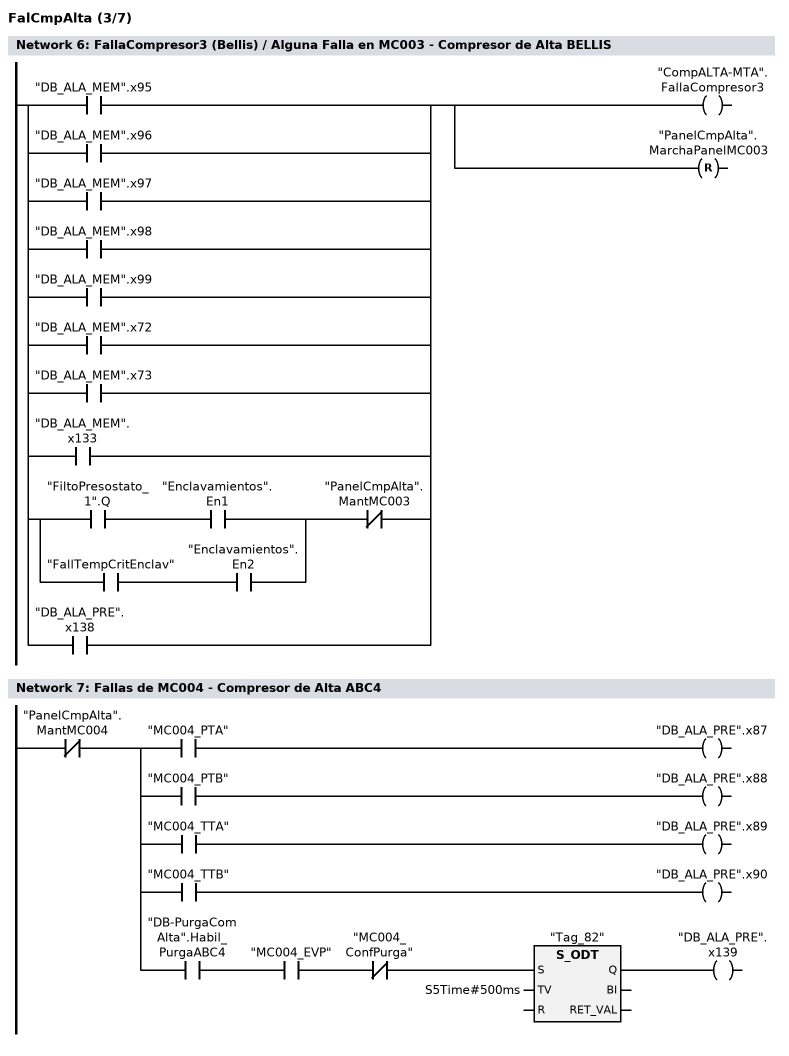
   RUNG wire#powerrail
      Contact( "DB_ALA_MEM".x95 )
      wire#w1
      Coil( "CompALTA-MTA".FallaCompresor3 )
   END_RUNG
   RUNG wire#powerrail
      Contact( "DB_ALA_MEM".x96 )
   END_RUNG wire#w1
   RUNG wire#powerrail
      Contact( "DB_ALA_MEM".x97 )
   END_RUNG wire#w1
   RUNG wire#powerrail
      Contact( "DB_ALA_MEM".x98 )
   END_RUNG wire#w1
   RUNG wire#powerrail
      Contact( "DB_ALA_MEM".x99 )
   END_RUNG wire#w1
   RUNG wire#powerrail
      Contact( "DB_ALA_MEM".x72 )
   END_RUNG wire#w1
   RUNG wire#powerrail
      Contact( "DB_ALA_MEM".x73 )
   END_RUNG wire#w1
   RUNG wire#powerrail
      Contact( "DB_ALA_MEM".x133 )
   END_RUNG wire#w1
   RUNG wire#powerrail
      Contact( "FiltoPresostato_1".Q )
      Contact( "Enclavamientos".En1 )
      wire#w2
      I_Contact( "PanelCmpAlta".MantMC003 )
   END_RUNG wire#w1
   RUNG wire#powerrail
      Contact( "FallTempCritEnclav" )
      Contact( "Enclavamientos".En2 )
   END_RUNG wire#w2
   RUNG wire#powerrail
      Contact( "DB_ALA_PRE".x138 )
   END_RUNG wire#w1
   RUNG wire#w1
      R_Coil( "PanelCmpAlta".MarchaPanelMC003 )
   END_RUNG
   // the same network as SCL:
   "CompALTA-MTA".FallaCompresor3 := "DB_ALA_MEM".x95 OR "DB_ALA_MEM".x96 OR "DB_ALA_MEM".x97 OR "DB_ALA_MEM".x98 OR "DB_ALA_MEM".x99 OR "DB_ALA_MEM".x72 OR "DB_ALA_MEM".x73 OR "DB_ALA_MEM".x133 OR ((("FiltoPresostato_1".Q AND "Enclavamientos".En1) OR ("FallTempCritEnclav" AND "Enclavamientos".En2)) AND NOT "PanelCmpAlta".MantMC003) OR "DB_ALA_PRE".x138;
   IF "CompALTA-MTA".FallaCompresor3 THEN "PanelCmpAlta".MarchaPanelMC003 := FALSE; END_IF;
END_REGION

REGION Network 7: Fallas de MC004 - Compresor de Alta ABC4
   RUNG wire#powerrail
      I_Contact( "PanelCmpAlta".MantMC004 )
      wire#w1
      Contact( "MC004_PTA" )
      Coil( "DB_ALA_PRE".x87 )
   END_RUNG
   RUNG wire#w1
      Contact( "MC004_PTB" )
      Coil( "DB_ALA_PRE".x88 )
   END_RUNG
   RUNG wire#w1
      Contact( "MC004_TTA" )
      Coil( "DB_ALA_PRE".x89 )
   END_RUNG
   RUNG wire#w1
      Contact( "MC004_TTB" )
      Coil( "DB_ALA_PRE".x90 )
   END_RUNG
   RUNG wire#w1
      Contact( "DB-PurgaComAlta".Habil_PurgaABC4 )
      Contact( "MC004_EVP" )
      I_Contact( "MC004_ConfPurga" )
      S_ODT(T_NO := "Tag_82", TV := S5Time#500ms, R :=, BI =>, RET_VAL =>)
      Coil( "DB_ALA_PRE".x139 )
   END_RUNG
   // the same network as SCL:
   #_w1 := NOT "PanelCmpAlta".MantMC004;
   "DB_ALA_PRE".x87 := #_w1 AND "MC004_PTA";
   "DB_ALA_PRE".x88 := #_w1 AND "MC004_PTB";
   "DB_ALA_PRE".x89 := #_w1 AND "MC004_TTA";
   "DB_ALA_PRE".x90 := #_w1 AND "MC004_TTB";
   #_s5time1 := S_ODT(T_NO := "Tag_82",
                      S := #_w1 AND "DB-PurgaComAlta".Habil_PurgaABC4 AND "MC004_EVP" AND NOT "MC004_ConfPurga",
                      TV := S5Time#500ms,
                      Q => #_w2);
   "DB_ALA_PRE".x139 := #_w2;
END_REGION

REGION Network 8: FallaCompresor4 (ABC4) / Alguna Falla en MC004 - Compresor de Alta ABC4
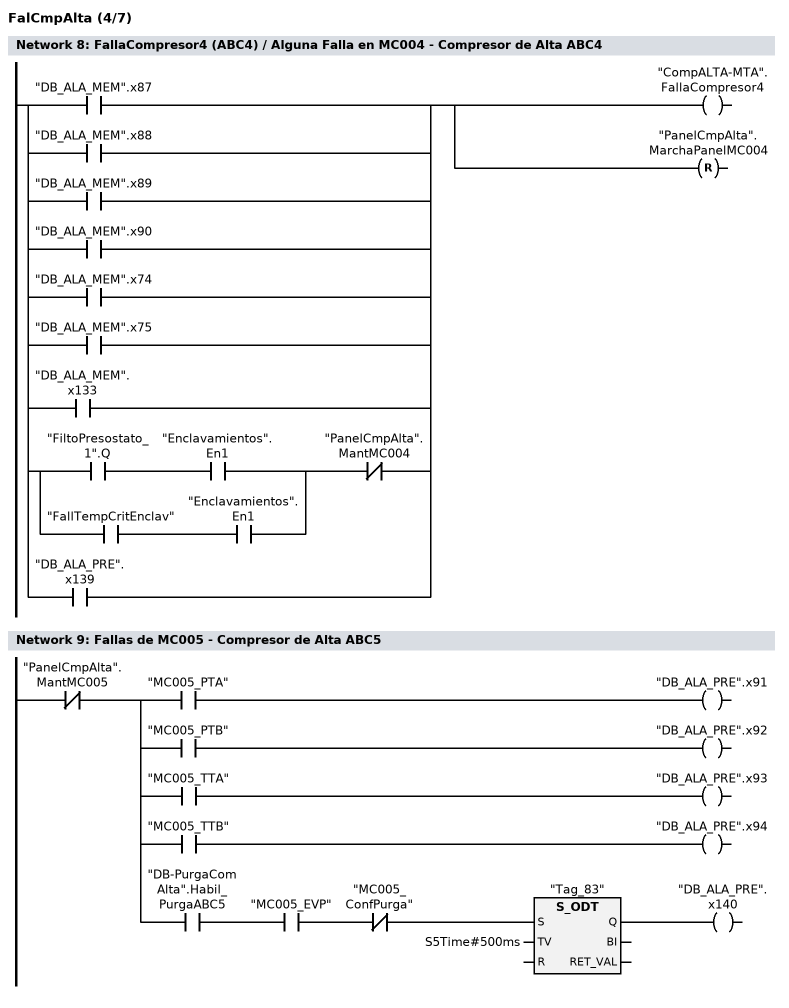
   RUNG wire#powerrail
      Contact( "DB_ALA_MEM".x87 )
      wire#w1
      Coil( "CompALTA-MTA".FallaCompresor4 )
   END_RUNG
   RUNG wire#powerrail
      Contact( "DB_ALA_MEM".x88 )
   END_RUNG wire#w1
   RUNG wire#powerrail
      Contact( "DB_ALA_MEM".x89 )
   END_RUNG wire#w1
   RUNG wire#powerrail
      Contact( "DB_ALA_MEM".x90 )
   END_RUNG wire#w1
   RUNG wire#powerrail
      Contact( "DB_ALA_MEM".x74 )
   END_RUNG wire#w1
   RUNG wire#powerrail
      Contact( "DB_ALA_MEM".x75 )
   END_RUNG wire#w1
   RUNG wire#powerrail
      Contact( "DB_ALA_MEM".x133 )
   END_RUNG wire#w1
   RUNG wire#powerrail
      Contact( "FiltoPresostato_1".Q )
      Contact( "Enclavamientos".En1 )
      wire#w2
      I_Contact( "PanelCmpAlta".MantMC004 )
   END_RUNG wire#w1
   RUNG wire#powerrail
      Contact( "FallTempCritEnclav" )
      Contact( "Enclavamientos".En1 )
   END_RUNG wire#w2
   RUNG wire#powerrail
      Contact( "DB_ALA_PRE".x139 )
   END_RUNG wire#w1
   RUNG wire#w1
      R_Coil( "PanelCmpAlta".MarchaPanelMC004 )
   END_RUNG
   // the same network as SCL:
   "CompALTA-MTA".FallaCompresor4 := "DB_ALA_MEM".x87 OR "DB_ALA_MEM".x88 OR "DB_ALA_MEM".x89 OR "DB_ALA_MEM".x90 OR "DB_ALA_MEM".x74 OR "DB_ALA_MEM".x75 OR "DB_ALA_MEM".x133 OR ((("FiltoPresostato_1".Q AND "Enclavamientos".En1) OR ("FallTempCritEnclav" AND "Enclavamientos".En1)) AND NOT "PanelCmpAlta".MantMC004) OR "DB_ALA_PRE".x139;
   IF "CompALTA-MTA".FallaCompresor4 THEN "PanelCmpAlta".MarchaPanelMC004 := FALSE; END_IF;
END_REGION

REGION Network 9: Fallas de MC005 - Compresor de Alta ABC5
   RUNG wire#powerrail
      I_Contact( "PanelCmpAlta".MantMC005 )
      wire#w1
      Contact( "MC005_PTA" )
      Coil( "DB_ALA_PRE".x91 )
   END_RUNG
   RUNG wire#w1
      Contact( "MC005_PTB" )
      Coil( "DB_ALA_PRE".x92 )
   END_RUNG
   RUNG wire#w1
      Contact( "MC005_TTA" )
      Coil( "DB_ALA_PRE".x93 )
   END_RUNG
   RUNG wire#w1
      Contact( "MC005_TTB" )
      Coil( "DB_ALA_PRE".x94 )
   END_RUNG
   RUNG wire#w1
      Contact( "DB-PurgaComAlta".Habil_PurgaABC5 )
      Contact( "MC005_EVP" )
      I_Contact( "MC005_ConfPurga" )
      S_ODT(T_NO := "Tag_83", TV := S5Time#500ms, R :=, BI =>, RET_VAL =>)
      Coil( "DB_ALA_PRE".x140 )
   END_RUNG
   // the same network as SCL:
   #_w1 := NOT "PanelCmpAlta".MantMC005;
   "DB_ALA_PRE".x91 := #_w1 AND "MC005_PTA";
   "DB_ALA_PRE".x92 := #_w1 AND "MC005_PTB";
   "DB_ALA_PRE".x93 := #_w1 AND "MC005_TTA";
   "DB_ALA_PRE".x94 := #_w1 AND "MC005_TTB";
   #_s5time1 := S_ODT(T_NO := "Tag_83",
                      S := #_w1 AND "DB-PurgaComAlta".Habil_PurgaABC5 AND "MC005_EVP" AND NOT "MC005_ConfPurga",
                      TV := S5Time#500ms,
                      Q => #_w2);
   "DB_ALA_PRE".x140 := #_w2;
END_REGION

REGION Network 10: FallaCompresor5 (ABC5) / Alguna Falla en MC005 - Compresor de Alta ABC5
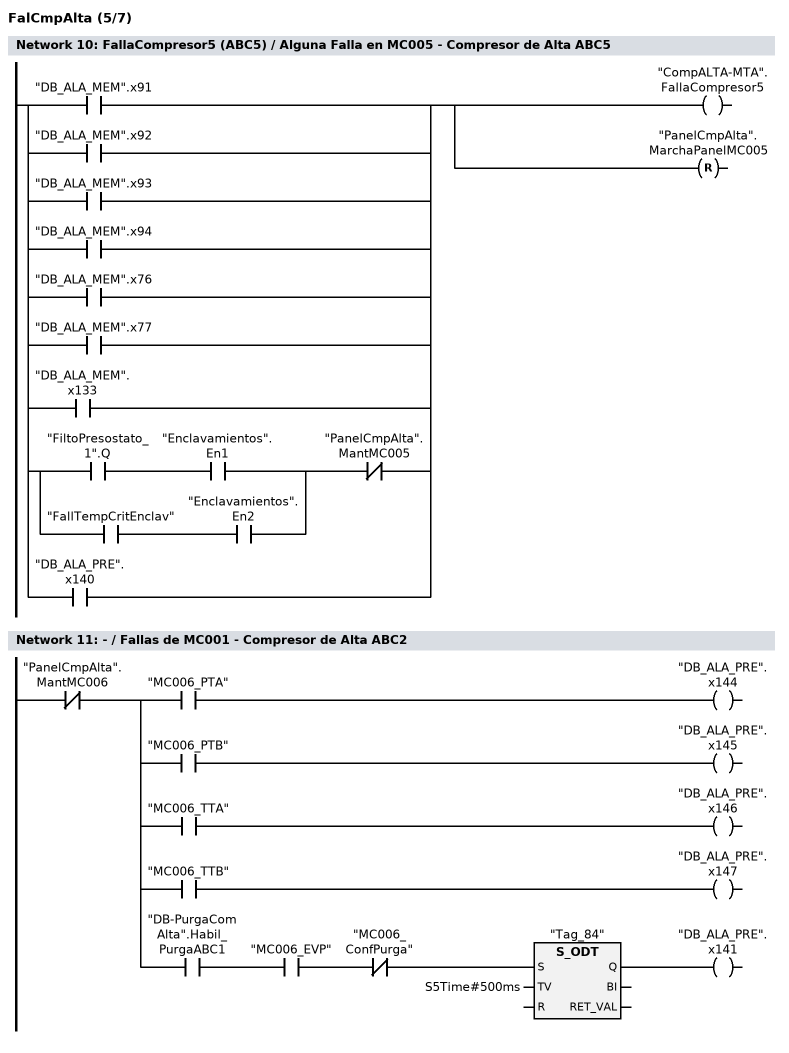
   RUNG wire#powerrail
      Contact( "DB_ALA_MEM".x91 )
      wire#w1
      Coil( "CompALTA-MTA".FallaCompresor5 )
   END_RUNG
   RUNG wire#powerrail
      Contact( "DB_ALA_MEM".x92 )
   END_RUNG wire#w1
   RUNG wire#powerrail
      Contact( "DB_ALA_MEM".x93 )
   END_RUNG wire#w1
   RUNG wire#powerrail
      Contact( "DB_ALA_MEM".x94 )
   END_RUNG wire#w1
   RUNG wire#powerrail
      Contact( "DB_ALA_MEM".x76 )
   END_RUNG wire#w1
   RUNG wire#powerrail
      Contact( "DB_ALA_MEM".x77 )
   END_RUNG wire#w1
   RUNG wire#powerrail
      Contact( "DB_ALA_MEM".x133 )
   END_RUNG wire#w1
   RUNG wire#powerrail
      Contact( "FiltoPresostato_1".Q )
      Contact( "Enclavamientos".En1 )
      wire#w2
      I_Contact( "PanelCmpAlta".MantMC005 )
   END_RUNG wire#w1
   RUNG wire#powerrail
      Contact( "FallTempCritEnclav" )
      Contact( "Enclavamientos".En2 )
   END_RUNG wire#w2
   RUNG wire#powerrail
      Contact( "DB_ALA_PRE".x140 )
   END_RUNG wire#w1
   RUNG wire#w1
      R_Coil( "PanelCmpAlta".MarchaPanelMC005 )
   END_RUNG
   // the same network as SCL:
   "CompALTA-MTA".FallaCompresor5 := "DB_ALA_MEM".x91 OR "DB_ALA_MEM".x92 OR "DB_ALA_MEM".x93 OR "DB_ALA_MEM".x94 OR "DB_ALA_MEM".x76 OR "DB_ALA_MEM".x77 OR "DB_ALA_MEM".x133 OR ((("FiltoPresostato_1".Q AND "Enclavamientos".En1) OR ("FallTempCritEnclav" AND "Enclavamientos".En2)) AND NOT "PanelCmpAlta".MantMC005) OR "DB_ALA_PRE".x140;
   IF "CompALTA-MTA".FallaCompresor5 THEN "PanelCmpAlta".MarchaPanelMC005 := FALSE; END_IF;
END_REGION

REGION Network 11: - / Fallas de MC001 - Compresor de Alta ABC2
   RUNG wire#powerrail
      I_Contact( "PanelCmpAlta".MantMC006 )
      wire#w1
      Contact( "MC006_PTA" )
      Coil( "DB_ALA_PRE".x144 )
   END_RUNG
   RUNG wire#w1
      Contact( "MC006_PTB" )
      Coil( "DB_ALA_PRE".x145 )
   END_RUNG
   RUNG wire#w1
      Contact( "MC006_TTA" )
      Coil( "DB_ALA_PRE".x146 )
   END_RUNG
   RUNG wire#w1
      Contact( "MC006_TTB" )
      Coil( "DB_ALA_PRE".x147 )
   END_RUNG
   RUNG wire#w1
      Contact( "DB-PurgaComAlta".Habil_PurgaABC1 )
      Contact( "MC006_EVP" )
      I_Contact( "MC006_ConfPurga" )
      S_ODT(T_NO := "Tag_84", TV := S5Time#500ms, R :=, BI =>, RET_VAL =>)
      Coil( "DB_ALA_PRE".x141 )
   END_RUNG
   // the same network as SCL:
   #_w1 := NOT "PanelCmpAlta".MantMC006;
   "DB_ALA_PRE".x144 := #_w1 AND "MC006_PTA";
   "DB_ALA_PRE".x145 := #_w1 AND "MC006_PTB";
   "DB_ALA_PRE".x146 := #_w1 AND "MC006_TTA";
   "DB_ALA_PRE".x147 := #_w1 AND "MC006_TTB";
   #_s5time1 := S_ODT(T_NO := "Tag_84",
                      S := #_w1 AND "DB-PurgaComAlta".Habil_PurgaABC1 AND "MC006_EVP" AND NOT "MC006_ConfPurga",
                      TV := S5Time#500ms,
                      Q => #_w2);
   "DB_ALA_PRE".x141 := #_w2;
END_REGION

REGION Network 12: FallaCompresor6 (ABC1) / Alguna Falla en MC001 - Compresor de Alta ABC2
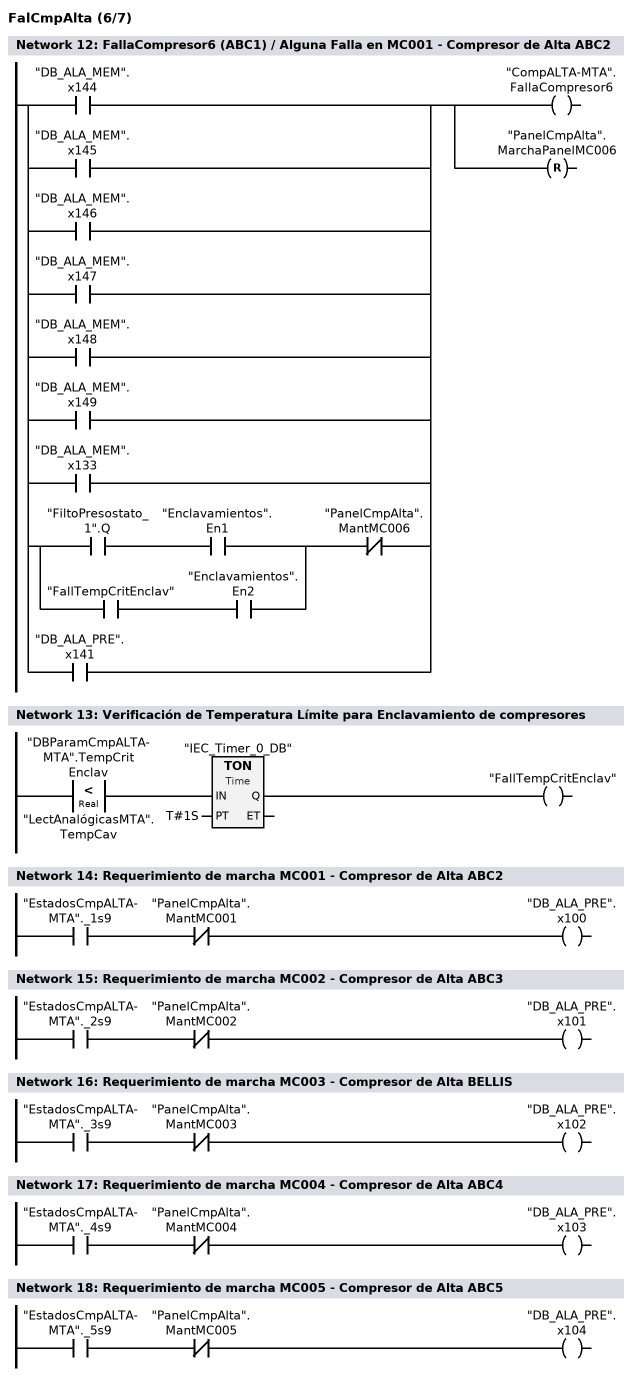
   RUNG wire#powerrail
      Contact( "DB_ALA_MEM".x144 )
      wire#w1
      Coil( "CompALTA-MTA".FallaCompresor6 )
   END_RUNG
   RUNG wire#powerrail
      Contact( "DB_ALA_MEM".x145 )
   END_RUNG wire#w1
   RUNG wire#powerrail
      Contact( "DB_ALA_MEM".x146 )
   END_RUNG wire#w1
   RUNG wire#powerrail
      Contact( "DB_ALA_MEM".x147 )
   END_RUNG wire#w1
   RUNG wire#powerrail
      Contact( "DB_ALA_MEM".x148 )
   END_RUNG wire#w1
   RUNG wire#powerrail
      Contact( "DB_ALA_MEM".x149 )
   END_RUNG wire#w1
   RUNG wire#powerrail
      Contact( "DB_ALA_MEM".x133 )
   END_RUNG wire#w1
   RUNG wire#powerrail
      Contact( "FiltoPresostato_1".Q )
      Contact( "Enclavamientos".En1 )
      wire#w2
      I_Contact( "PanelCmpAlta".MantMC006 )
   END_RUNG wire#w1
   RUNG wire#powerrail
      Contact( "FallTempCritEnclav" )
      Contact( "Enclavamientos".En2 )
   END_RUNG wire#w2
   RUNG wire#powerrail
      Contact( "DB_ALA_PRE".x141 )
   END_RUNG wire#w1
   RUNG wire#w1
      R_Coil( "PanelCmpAlta".MarchaPanelMC006 )
   END_RUNG
   // the same network as SCL:
   "CompALTA-MTA".FallaCompresor6 := "DB_ALA_MEM".x144 OR "DB_ALA_MEM".x145 OR "DB_ALA_MEM".x146 OR "DB_ALA_MEM".x147 OR "DB_ALA_MEM".x148 OR "DB_ALA_MEM".x149 OR "DB_ALA_MEM".x133 OR ((("FiltoPresostato_1".Q AND "Enclavamientos".En1) OR ("FallTempCritEnclav" AND "Enclavamientos".En2)) AND NOT "PanelCmpAlta".MantMC006) OR "DB_ALA_PRE".x141;
   IF "CompALTA-MTA".FallaCompresor6 THEN "PanelCmpAlta".MarchaPanelMC006 := FALSE; END_IF;
END_REGION

REGION Network 13: Verificación de Temperatura Límite para Enclavamiento de compresores
   "IEC_Timer_0_DB".TON(IN := "DBParamCmpALTA-MTA".TempCritEnclav < "LectAnalógicasMTA".TempCav, PT := T#1S);
   "FallTempCritEnclav" := "IEC_Timer_0_DB".Q;
END_REGION

REGION Network 14: Requerimiento de marcha MC001 - Compresor de Alta ABC2
   RUNG wire#powerrail
      Contact( "EstadosCmpALTA-MTA"._1s9 )
      I_Contact( "PanelCmpAlta".MantMC001 )
      Coil( "DB_ALA_PRE".x100 )
   END_RUNG
   // the same network as SCL:
   "DB_ALA_PRE".x100 := "EstadosCmpALTA-MTA"._1s9 AND NOT "PanelCmpAlta".MantMC001;
END_REGION

REGION Network 15: Requerimiento de marcha MC002 - Compresor de Alta ABC3
   RUNG wire#powerrail
      Contact( "EstadosCmpALTA-MTA"._2s9 )
      I_Contact( "PanelCmpAlta".MantMC002 )
      Coil( "DB_ALA_PRE".x101 )
   END_RUNG
   // the same network as SCL:
   "DB_ALA_PRE".x101 := "EstadosCmpALTA-MTA"._2s9 AND NOT "PanelCmpAlta".MantMC002;
END_REGION

REGION Network 16: Requerimiento de marcha MC003 - Compresor de Alta BELLIS
   RUNG wire#powerrail
      Contact( "EstadosCmpALTA-MTA"._3s9 )
      I_Contact( "PanelCmpAlta".MantMC003 )
      Coil( "DB_ALA_PRE".x102 )
   END_RUNG
   // the same network as SCL:
   "DB_ALA_PRE".x102 := "EstadosCmpALTA-MTA"._3s9 AND NOT "PanelCmpAlta".MantMC003;
END_REGION

REGION Network 17: Requerimiento de marcha MC004 - Compresor de Alta ABC4
   RUNG wire#powerrail
      Contact( "EstadosCmpALTA-MTA"._4s9 )
      I_Contact( "PanelCmpAlta".MantMC004 )
      Coil( "DB_ALA_PRE".x103 )
   END_RUNG
   // the same network as SCL:
   "DB_ALA_PRE".x103 := "EstadosCmpALTA-MTA"._4s9 AND NOT "PanelCmpAlta".MantMC004;
END_REGION

REGION Network 18: Requerimiento de marcha MC005 - Compresor de Alta ABC5
   RUNG wire#powerrail
      Contact( "EstadosCmpALTA-MTA"._5s9 )
      I_Contact( "PanelCmpAlta".MantMC005 )
      Coil( "DB_ALA_PRE".x104 )
   END_RUNG
   // the same network as SCL:
   "DB_ALA_PRE".x104 := "EstadosCmpALTA-MTA"._5s9 AND NOT "PanelCmpAlta".MantMC005;
END_REGION

REGION Network 19: Requerimiento de marcha MC001 - Compresor de Alta ABC2
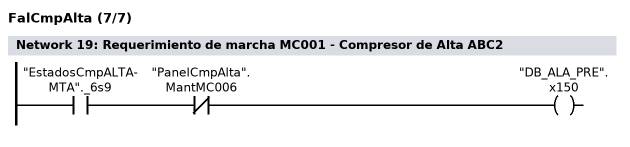
   RUNG wire#powerrail
      Contact( "EstadosCmpALTA-MTA"._6s9 )
      I_Contact( "PanelCmpAlta".MantMC006 )
      Coil( "DB_ALA_PRE".x150 )
   END_RUNG
   // the same network as SCL:
   "DB_ALA_PRE".x150 := "EstadosCmpALTA-MTA"._6s9 AND NOT "PanelCmpAlta".MantMC006;
END_REGION
END_FUNCTION

// folder: Auxiliares

FUNCTION "AjusteEntrada-SalidaMTA" : Void   // FC6, LAD
{ S7_Optimized_Access := 'FALSE' }
VERSION : 0.1
BEGIN

REGION Network 1
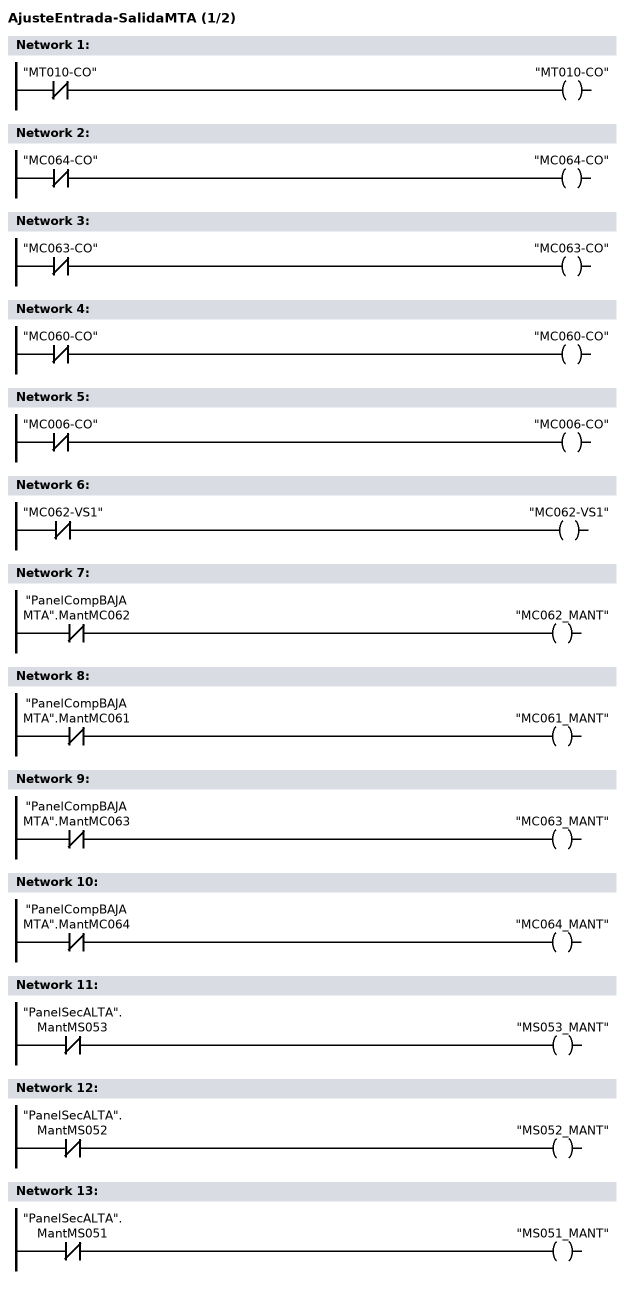
   RUNG wire#powerrail
      I_Contact( "MT010-CO" )
      Coil( "MT010-CO" )
   END_RUNG
   // the same network as SCL:
   "MT010-CO" := NOT "MT010-CO";
END_REGION

REGION Network 2
   RUNG wire#powerrail
      I_Contact( "MC064-CO" )
      Coil( "MC064-CO" )
   END_RUNG
   // the same network as SCL:
   "MC064-CO" := NOT "MC064-CO";
END_REGION

REGION Network 3
   RUNG wire#powerrail
      I_Contact( "MC063-CO" )
      Coil( "MC063-CO" )
   END_RUNG
   // the same network as SCL:
   "MC063-CO" := NOT "MC063-CO";
END_REGION

REGION Network 4
   RUNG wire#powerrail
      I_Contact( "MC060-CO" )
      Coil( "MC060-CO" )
   END_RUNG
   // the same network as SCL:
   "MC060-CO" := NOT "MC060-CO";
END_REGION

REGION Network 5
   RUNG wire#powerrail
      I_Contact( "MC006-CO" )
      Coil( "MC006-CO" )
   END_RUNG
   // the same network as SCL:
   "MC006-CO" := NOT "MC006-CO";
END_REGION

REGION Network 6
   RUNG wire#powerrail
      I_Contact( "MC062-VS1" )
      Coil( "MC062-VS1" )
   END_RUNG
   // the same network as SCL:
   "MC062-VS1" := NOT "MC062-VS1";
END_REGION

REGION Network 7
   RUNG wire#powerrail
      I_Contact( "PanelCompBAJA MTA".MantMC062 )
      Coil( "MC062_MANT" )
   END_RUNG
   // the same network as SCL:
   "MC062_MANT" := NOT "PanelCompBAJA MTA".MantMC062;
END_REGION

REGION Network 8
   RUNG wire#powerrail
      I_Contact( "PanelCompBAJA MTA".MantMC061 )
      Coil( "MC061_MANT" )
   END_RUNG
   // the same network as SCL:
   "MC061_MANT" := NOT "PanelCompBAJA MTA".MantMC061;
END_REGION

REGION Network 9
   RUNG wire#powerrail
      I_Contact( "PanelCompBAJA MTA".MantMC063 )
      Coil( "MC063_MANT" )
   END_RUNG
   // the same network as SCL:
   "MC063_MANT" := NOT "PanelCompBAJA MTA".MantMC063;
END_REGION

REGION Network 10
   RUNG wire#powerrail
      I_Contact( "PanelCompBAJA MTA".MantMC064 )
      Coil( "MC064_MANT" )
   END_RUNG
   // the same network as SCL:
   "MC064_MANT" := NOT "PanelCompBAJA MTA".MantMC064;
END_REGION

REGION Network 11
   RUNG wire#powerrail
      I_Contact( "PanelSecALTA".MantMS053 )
      Coil( "MS053_MANT" )
   END_RUNG
   // the same network as SCL:
   "MS053_MANT" := NOT "PanelSecALTA".MantMS053;
END_REGION

REGION Network 12
   RUNG wire#powerrail
      I_Contact( "PanelSecALTA".MantMS052 )
      Coil( "MS052_MANT" )
   END_RUNG
   // the same network as SCL:
   "MS052_MANT" := NOT "PanelSecALTA".MantMS052;
END_REGION

REGION Network 13
   RUNG wire#powerrail
      I_Contact( "PanelSecALTA".MantMS051 )
      Coil( "MS051_MANT" )
   END_RUNG
   // the same network as SCL:
   "MS051_MANT" := NOT "PanelSecALTA".MantMS051;
END_REGION

REGION Network 14
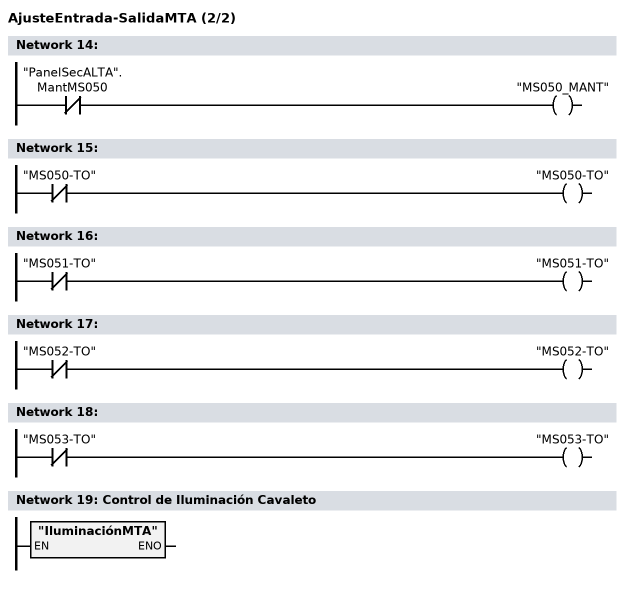
   RUNG wire#powerrail
      I_Contact( "PanelSecALTA".MantMS050 )
      Coil( "MS050_MANT" )
   END_RUNG
   // the same network as SCL:
   "MS050_MANT" := NOT "PanelSecALTA".MantMS050;
END_REGION

REGION Network 15
   RUNG wire#powerrail
      I_Contact( "MS050-TO" )
      Coil( "MS050-TO" )
   END_RUNG
   // the same network as SCL:
   "MS050-TO" := NOT "MS050-TO";
END_REGION

REGION Network 16
   RUNG wire#powerrail
      I_Contact( "MS051-TO" )
      Coil( "MS051-TO" )
   END_RUNG
   // the same network as SCL:
   "MS051-TO" := NOT "MS051-TO";
END_REGION

REGION Network 17
   RUNG wire#powerrail
      I_Contact( "MS052-TO" )
      Coil( "MS052-TO" )
   END_RUNG
   // the same network as SCL:
   "MS052-TO" := NOT "MS052-TO";
END_REGION

REGION Network 18
   RUNG wire#powerrail
      I_Contact( "MS053-TO" )
      Coil( "MS053-TO" )
   END_RUNG
   // the same network as SCL:
   "MS053-TO" := NOT "MS053-TO";
END_REGION

REGION Network 19: Control de Iluminación Cavaleto
   RUNG wire#powerrail
      "IluminaciónMTA"()
   END_RUNG
   // the same network as SCL:
   "IluminaciónMTA"();
END_REGION
END_FUNCTION

FUNCTION "And-Byte MTA" : Void   // FC22, LAD
{ S7_Optimized_Access := 'FALSE' }
VERSION : 0.1
BEGIN

REGION Network 1
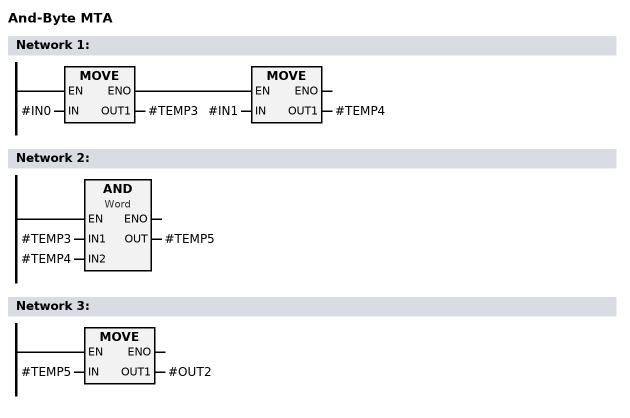
   RUNG wire#powerrail
      { S7_GenerateENO := "TRUE" } Move(in := #IN0, out1 => #TEMP3)
      { S7_GenerateENO := "TRUE" } Move(in := #IN1, out1 => #TEMP4)
   END_RUNG
   // the same network as SCL:
   // ENO of a box is taken as its EN; it also drops when the box reports an error
   #TEMP3 := #IN0;
   #TEMP4 := #IN1;
END_REGION

REGION Network 2
   RUNG wire#powerrail
      { S7_Templates := "SrcType := Word"; S7_GenerateENO := "TRUE" } And(in1 := #TEMP3, in2 := #TEMP4, out => #TEMP5)
   END_RUNG
   // the same network as SCL:
   #TEMP5 := #TEMP3 AND #TEMP4;
END_REGION

REGION Network 3
   RUNG wire#powerrail
      { S7_GenerateENO := "TRUE" } Move(in := #TEMP5, out1 => #OUT2)
   END_RUNG
   // the same network as SCL:
   #OUT2 := #TEMP5;
END_REGION
END_FUNCTION

FUNCTION "Inicialización" : Void   // FC46, LAD
{ S7_Optimized_Access := 'FALSE' }
VERSION : 0.1
BEGIN

REGION Network 1
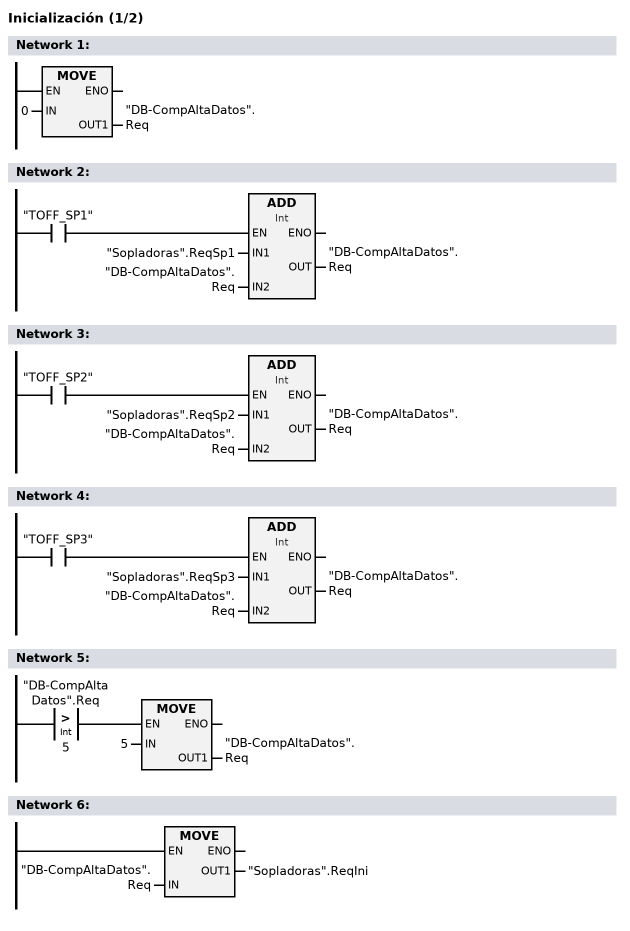
   RUNG wire#powerrail
      { S7_GenerateENO := "TRUE" } Move(in := 0, out1 => "DB-CompAltaDatos".Req)
   END_RUNG
   // the same network as SCL:
   "DB-CompAltaDatos".Req := 0;
END_REGION

REGION Network 2
   RUNG wire#powerrail
      Contact( "TOFF_SP1" )
      { S7_Templates := "SrcType := Int"; S7_GenerateENO := "TRUE" } Add(in1 := "Sopladoras".ReqSp1, in2 := "DB-CompAltaDatos".Req, out => "DB-CompAltaDatos".Req)
   END_RUNG
   // the same network as SCL:
   IF "TOFF_SP1" THEN "DB-CompAltaDatos".Req := "Sopladoras".ReqSp1 + "DB-CompAltaDatos".Req; END_IF;
END_REGION

REGION Network 3
   RUNG wire#powerrail
      Contact( "TOFF_SP2" )
      { S7_Templates := "SrcType := Int"; S7_GenerateENO := "TRUE" } Add(in1 := "Sopladoras".ReqSp2, in2 := "DB-CompAltaDatos".Req, out => "DB-CompAltaDatos".Req)
   END_RUNG
   // the same network as SCL:
   IF "TOFF_SP2" THEN "DB-CompAltaDatos".Req := "Sopladoras".ReqSp2 + "DB-CompAltaDatos".Req; END_IF;
END_REGION

REGION Network 4
   RUNG wire#powerrail
      Contact( "TOFF_SP3" )
      { S7_Templates := "SrcType := Int"; S7_GenerateENO := "TRUE" } Add(in1 := "Sopladoras".ReqSp3, in2 := "DB-CompAltaDatos".Req, out => "DB-CompAltaDatos".Req)
   END_RUNG
   // the same network as SCL:
   IF "TOFF_SP3" THEN "DB-CompAltaDatos".Req := "Sopladoras".ReqSp3 + "DB-CompAltaDatos".Req; END_IF;
END_REGION

REGION Network 5
   RUNG wire#powerrail
      { S7_Templates := "SrcType := Int" } GT_Contact(in1 := "DB-CompAltaDatos".Req, in2 := 5)
      { S7_GenerateENO := "TRUE" } Move(in := 5, out1 => "DB-CompAltaDatos".Req)
   END_RUNG
   // the same network as SCL:
   IF "DB-CompAltaDatos".Req > 5 THEN "DB-CompAltaDatos".Req := 5; END_IF;
END_REGION

REGION Network 6
   RUNG wire#powerrail
      { S7_GenerateENO := "TRUE" } Move(in := "DB-CompAltaDatos".Req, out1 => "Sopladoras".ReqIni)
   END_RUNG
   // the same network as SCL:
   "Sopladoras".ReqIni := "DB-CompAltaDatos".Req;
END_REGION

REGION Network 7
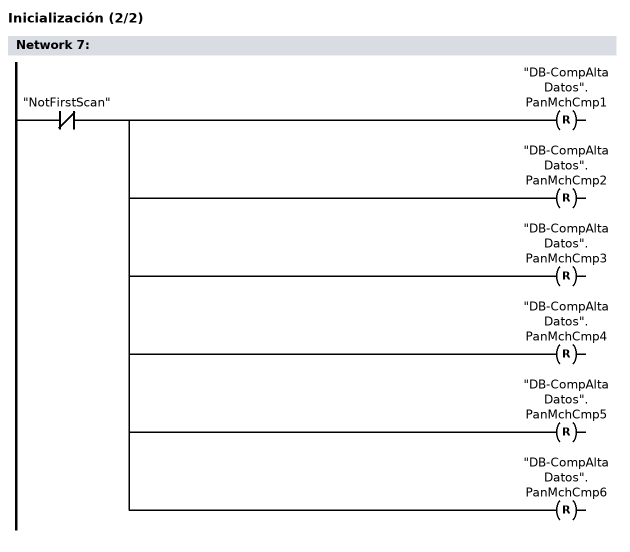
   RUNG wire#powerrail
      I_Contact( "NotFirstScan" )
      wire#w1
      R_Coil( "DB-CompAltaDatos".PanMchCmp1 )
   END_RUNG
   RUNG wire#w1
      R_Coil( "DB-CompAltaDatos".PanMchCmp2 )
   END_RUNG
   RUNG wire#w1
      R_Coil( "DB-CompAltaDatos".PanMchCmp3 )
   END_RUNG
   RUNG wire#w1
      R_Coil( "DB-CompAltaDatos".PanMchCmp4 )
   END_RUNG
   RUNG wire#w1
      R_Coil( "DB-CompAltaDatos".PanMchCmp5 )
   END_RUNG
   RUNG wire#w1
      R_Coil( "DB-CompAltaDatos".PanMchCmp6 )
   END_RUNG
   // the same network as SCL:
   IF NOT "NotFirstScan" THEN
       "DB-CompAltaDatos".PanMchCmp1 := FALSE;
       "DB-CompAltaDatos".PanMchCmp2 := FALSE;
       "DB-CompAltaDatos".PanMchCmp3 := FALSE;
       "DB-CompAltaDatos".PanMchCmp4 := FALSE;
       "DB-CompAltaDatos".PanMchCmp5 := FALSE;
       "DB-CompAltaDatos".PanMchCmp6 := FALSE;
   END_IF;
END_REGION
END_FUNCTION

// folder: Bloques Estándar

FUNCTION_BLOCK "ControladorMotoresMTA"   // FB2, LAD
{ S7_Optimized_Access := 'FALSE' }
VERSION : 0.1
BEGIN

REGION Network 2
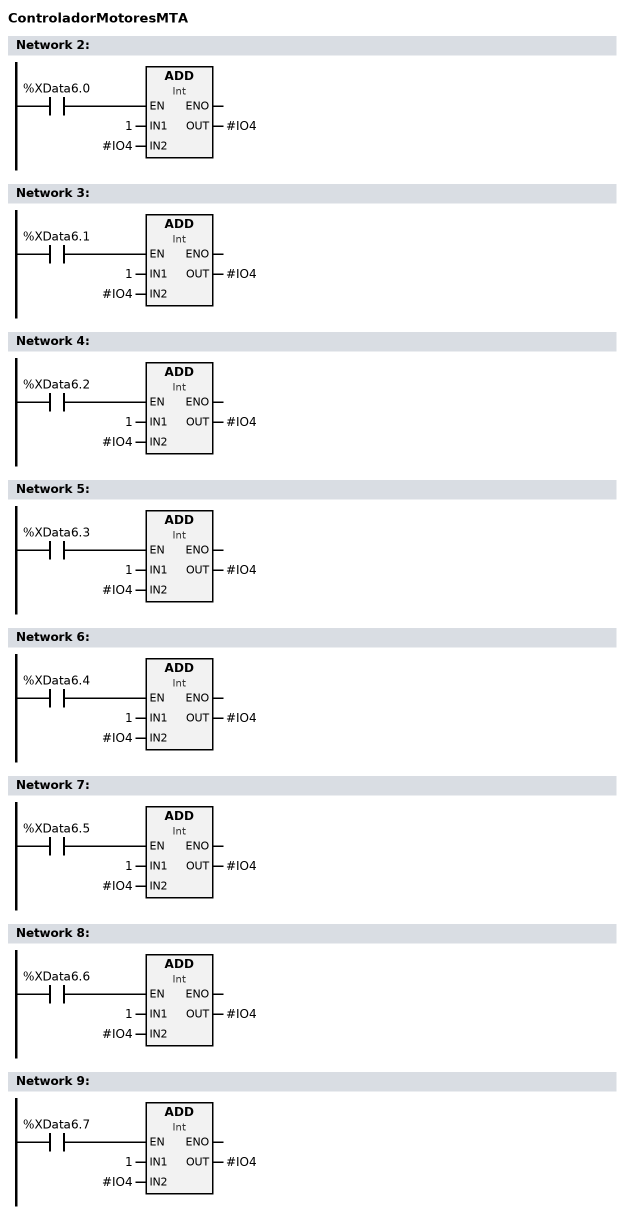
   RUNG wire#powerrail
      Contact( %XData6.0 )
      { S7_Templates := "SrcType := Int"; S7_GenerateENO := "TRUE" } Add(in1 := 1, in2 := #IO4, out => #IO4)
   END_RUNG
   // the same network as SCL:
   IF %XData6.0 THEN #IO4 := 1 + #IO4; END_IF;
END_REGION

REGION Network 3
   RUNG wire#powerrail
      Contact( %XData6.1 )
      { S7_Templates := "SrcType := Int"; S7_GenerateENO := "TRUE" } Add(in1 := 1, in2 := #IO4, out => #IO4)
   END_RUNG
   // the same network as SCL:
   IF %XData6.1 THEN #IO4 := 1 + #IO4; END_IF;
END_REGION

REGION Network 4
   RUNG wire#powerrail
      Contact( %XData6.2 )
      { S7_Templates := "SrcType := Int"; S7_GenerateENO := "TRUE" } Add(in1 := 1, in2 := #IO4, out => #IO4)
   END_RUNG
   // the same network as SCL:
   IF %XData6.2 THEN #IO4 := 1 + #IO4; END_IF;
END_REGION

REGION Network 5
   RUNG wire#powerrail
      Contact( %XData6.3 )
      { S7_Templates := "SrcType := Int"; S7_GenerateENO := "TRUE" } Add(in1 := 1, in2 := #IO4, out => #IO4)
   END_RUNG
   // the same network as SCL:
   IF %XData6.3 THEN #IO4 := 1 + #IO4; END_IF;
END_REGION

REGION Network 6
   RUNG wire#powerrail
      Contact( %XData6.4 )
      { S7_Templates := "SrcType := Int"; S7_GenerateENO := "TRUE" } Add(in1 := 1, in2 := #IO4, out => #IO4)
   END_RUNG
   // the same network as SCL:
   IF %XData6.4 THEN #IO4 := 1 + #IO4; END_IF;
END_REGION

REGION Network 7
   RUNG wire#powerrail
      Contact( %XData6.5 )
      { S7_Templates := "SrcType := Int"; S7_GenerateENO := "TRUE" } Add(in1 := 1, in2 := #IO4, out => #IO4)
   END_RUNG
   // the same network as SCL:
   IF %XData6.5 THEN #IO4 := 1 + #IO4; END_IF;
END_REGION

REGION Network 8
   RUNG wire#powerrail
      Contact( %XData6.6 )
      { S7_Templates := "SrcType := Int"; S7_GenerateENO := "TRUE" } Add(in1 := 1, in2 := #IO4, out => #IO4)
   END_RUNG
   // the same network as SCL:
   IF %XData6.6 THEN #IO4 := 1 + #IO4; END_IF;
END_REGION

REGION Network 9
   RUNG wire#powerrail
      Contact( %XData6.7 )
      { S7_Templates := "SrcType := Int"; S7_GenerateENO := "TRUE" } Add(in1 := 1, in2 := #IO4, out => #IO4)
   END_RUNG
   // the same network as SCL:
   IF %XData6.7 THEN #IO4 := 1 + #IO4; END_IF;
END_REGION
END_FUNCTION_BLOCK

// folder: Compresores/Alta

FUNCTION "CompresoresAltaMTA" : Void   // FC13, LAD
{ S7_Optimized_Access := 'FALSE' }
VERSION : 0.1
BEGIN

REGION Network 1
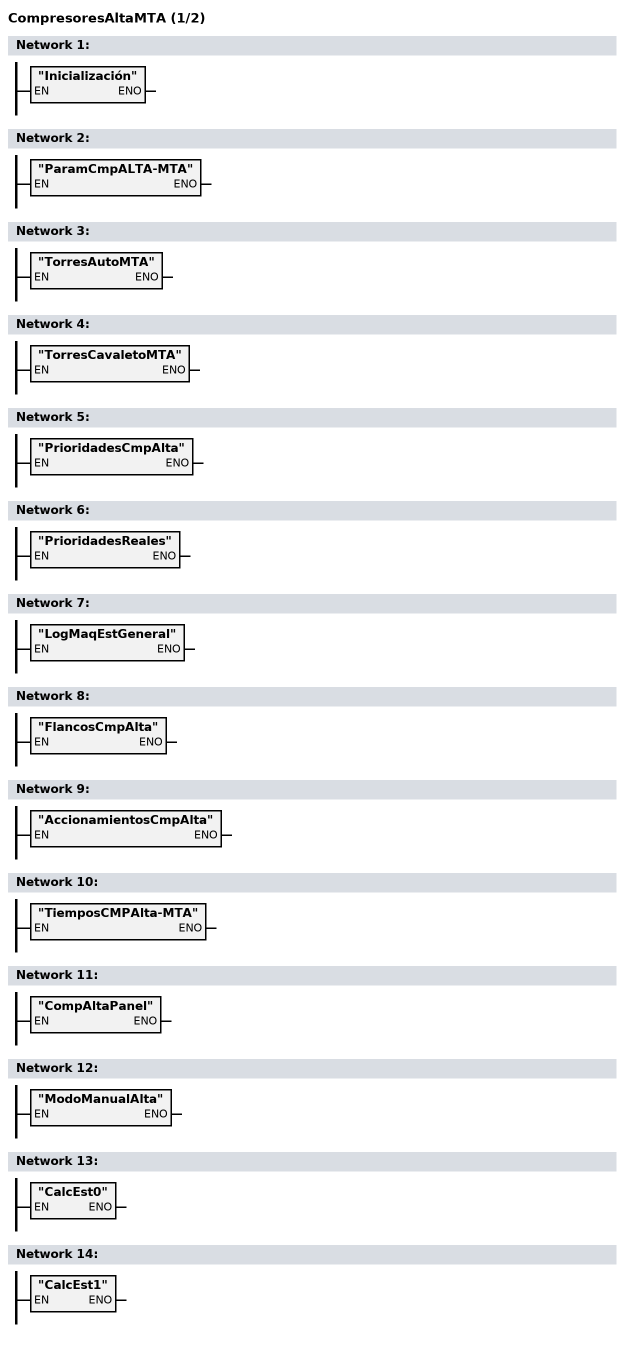
   RUNG wire#powerrail
      "Inicialización"()
   END_RUNG
   // the same network as SCL:
   "Inicialización"();
END_REGION

REGION Network 2
   RUNG wire#powerrail
      "ParamCmpALTA-MTA"()
   END_RUNG
   // the same network as SCL:
   "ParamCmpALTA-MTA"();
END_REGION

REGION Network 3
   RUNG wire#powerrail
      "TorresAutoMTA"()
   END_RUNG
   // the same network as SCL:
   "TorresAutoMTA"();
END_REGION

REGION Network 4
   RUNG wire#powerrail
      "TorresCavaletoMTA"()
   END_RUNG
   // the same network as SCL:
   "TorresCavaletoMTA"();
END_REGION

REGION Network 5
   RUNG wire#powerrail
      "PrioridadesCmpAlta"()
   END_RUNG
   // the same network as SCL:
   "PrioridadesCmpAlta"();
END_REGION

REGION Network 6
   RUNG wire#powerrail
      "PrioridadesReales"()
   END_RUNG
   // the same network as SCL:
   "PrioridadesReales"();
END_REGION

REGION Network 7
   RUNG wire#powerrail
      "LogMaqEstGeneral"()
   END_RUNG
   // the same network as SCL:
   "LogMaqEstGeneral"();
END_REGION

REGION Network 8
   RUNG wire#powerrail
      "FlancosCmpAlta"()
   END_RUNG
   // the same network as SCL:
   "FlancosCmpAlta"();
END_REGION

REGION Network 9
   RUNG wire#powerrail
      "AccionamientosCmpAlta"()
   END_RUNG
   // the same network as SCL:
   "AccionamientosCmpAlta"();
END_REGION

REGION Network 10
   RUNG wire#powerrail
      "TiemposCMPAlta-MTA"()
   END_RUNG
   // the same network as SCL:
   "TiemposCMPAlta-MTA"();
END_REGION

REGION Network 11
   RUNG wire#powerrail
      "CompAltaPanel"()
   END_RUNG
   // the same network as SCL:
   "CompAltaPanel"();
END_REGION

REGION Network 12
   RUNG wire#powerrail
      "ModoManualAlta"()
   END_RUNG
   // the same network as SCL:
   "ModoManualAlta"();
END_REGION

REGION Network 13
   RUNG wire#powerrail
      "CalcEst0"()
   END_RUNG
   // the same network as SCL:
   "CalcEst0"();
END_REGION

REGION Network 14
   RUNG wire#powerrail
      "CalcEst1"()
   END_RUNG
   // the same network as SCL:
   "CalcEst1"();
END_REGION

REGION Network 15
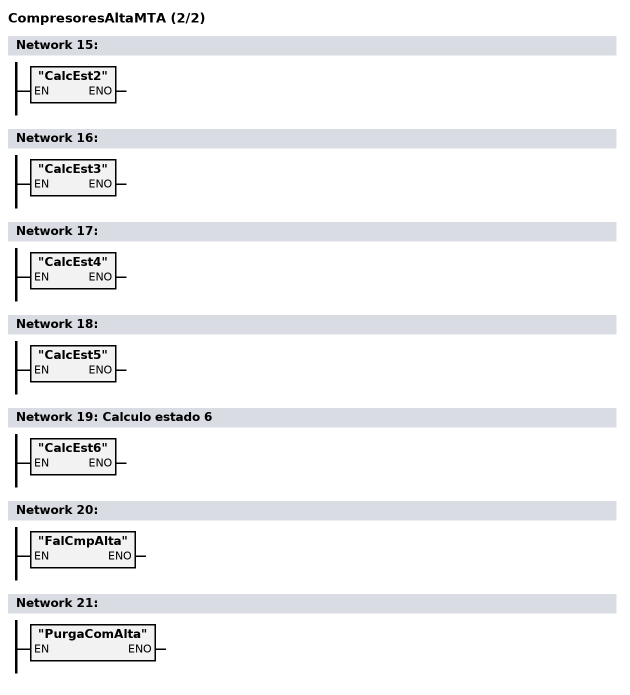
   RUNG wire#powerrail
      "CalcEst2"()
   END_RUNG
   // the same network as SCL:
   "CalcEst2"();
END_REGION

REGION Network 16
   RUNG wire#powerrail
      "CalcEst3"()
   END_RUNG
   // the same network as SCL:
   "CalcEst3"();
END_REGION

REGION Network 17
   RUNG wire#powerrail
      "CalcEst4"()
   END_RUNG
   // the same network as SCL:
   "CalcEst4"();
END_REGION

REGION Network 18
   RUNG wire#powerrail
      "CalcEst5"()
   END_RUNG
   // the same network as SCL:
   "CalcEst5"();
END_REGION

REGION Network 19: Calculo estado 6
   RUNG wire#powerrail
      "CalcEst6"()
   END_RUNG
   // the same network as SCL:
   "CalcEst6"();
END_REGION

REGION Network 20
   RUNG wire#powerrail
      "FalCmpAlta"()
   END_RUNG
   // the same network as SCL:
   "FalCmpAlta"();
END_REGION

REGION Network 21
   RUNG wire#powerrail
      "PurgaComAlta"()
   END_RUNG
   // the same network as SCL:
   "PurgaComAlta"();
END_REGION
END_FUNCTION

FUNCTION "ParamCmpALTA-MTA" : Void   // FC30, LAD
{ S7_Optimized_Access := 'FALSE' }
VERSION : 0.1
BEGIN

REGION Network 1
